TYPE "UDT012_Recirculation"
TITLE = State of recirculation mode
VERSION : 0.0
   STRUCT
      Intervall : Bool;   // Recirculation in interval mode (reduced or low pressure circulation)
      Parallel : Bool;   // Parallel circulation is activ (not used)
      Lowpressure : Bool;   // Low pressure circulation is active
      Reduced : Bool;   // Reduced circulation is active
      Highpressure : Bool;   // High pressure circulation over one mixing head is active
      Tolerance_OK : Bool;   // Request wether tolarances of the analog values at PUC are OK
      Weekendswitching : Bool;   // The pouring machine is in weekend mode
      Pausetime : Bool;   // The pouring machine is pausing time of the interval
      Break_KK : Bool;   // Stop flag of a active circulation mode to fill cylinder of a cylinder machine
      HP_is_active : Bool;   // High pressure circulation is active
      Is_selected : Bool;   // A circulation mode of the pouring machine is selected
      RequestPausePos : Bool;   // Request to the cylinder machine to bring the cylinder in break position
      cycle_runs : Bool;   // Save flag of the stop flag while starting a pouring cycle
      Is_active : Bool;   // A cycle mode of the pouring machine is active (no fault and oparition mode OK)
      Lowpressure_Exist : Bool;   // Low pressure circulation is existing
      Spare_1_7 : Bool;
      Switch_Intervall : Bool;   // Switch circulation in interval mode (reduced or low pressure circulation) selected
      Switch_Parallel : Bool;   // Switch Parallel circulation is selected (not used)
      Switch_Lowpressure : Bool;   // Switch Low pressure circulation is selected
      Switch_Reduced : Bool;   // Switch Reduced circulation is selected
      Intervall_Reduced : Bool;   // Reduced circulation in Intervall is active
      Intervall_Lowpressure : Bool;   // Low pressure circulation in Intervall is active
      Intervall_Reduced_Pause : Bool;   // Reduced circulation in Intervall pause is active
      Intervall_Lowpressure_Pause : Bool;   // Low pressure circulation in Intervall pause is active
      Spare_3_0 : Bool;
      Spare_3_1 : Bool;
      Spare_3_2 : Bool;
      Spare_3_3 : Bool;
      Spare_3_4 : Bool;
      Spare_3_5 : Bool;
      Spare_3_6 : Bool;
      Spare_3_7 : Bool;
      State_Intervall : Int;
      State_Lowpressure : Int;
      State_Reduced : Int;
      Indicator_HP : "UDT001_DWord_1_32";   // Indicates selected high pressure circulation
      Status_RC_HP : Int;   // Flag of the steps select and deselect high pressure circulation
      Button_HP : "UDT001_DWord_1_32";   // Button to select high pressure circulation
      Lamp_HP : "UDT001_DWord_1_32";   // Activation of lamps to indicat that high pressure recirculation runs
      SWU_RC_HP : DWord;   // Bitvalue of the SWU-Number where high pressure circulation runs
   END_STRUCT;
END_TYPE

TYPE "UDT013_Robot"
VERSION : 0.1
   STRUCT
      Switches : Struct
         SwitchHomePosON_OFF : Bool;   // Switch home position on/off
         SwitchMaintPosON_OFF : Bool;   // Switch maintenance position on/off
         SwitchTestShotON_OFF : Bool;   // Switch to make a couple shot with roboter
         SwitchCleaningON_OFF : Bool;   // Switch cleaning program on/off
         SwitchBrushON_OFF : Bool;   // Switch brush program on/off
         SwitchSyncON_OFF : Bool;   // Switch for checking EPS
         SwitchEnableRobotON_OFF : Bool;   // Switch no foaming in the conveyor (conveyor standalone)
         SwitchLearningON_OFF : Bool;   // Switch for learning the shot path (in conection with Shotware)
         SwitchTeachingON_OFF : Bool;   // Switch for Teaching the Robot
         Switch_10 : Bool;
         Switch_11 : Bool;
         Switch_12 : Bool;
         Switch_13 : Bool;
         Switch_14 : Bool;
         Switch_15 : Bool;
         Switch_16 : Bool;
         StateHomePos : Byte;   // 1->Drive ON; 2->Fault Drive; 3->Drive requested but not on
         StateMaintPos : Byte;   // 1->Drive ON; 2->Fault Drive; 3->Drive requested but not on
         StateTestShot : Byte;   // 1->Drive ON; 2->Fault Drive; 3->Drive requested but not on
         StateCleaning : Byte;   // 1->Drive ON; 2->Fault Drive; 3->Drive requested but not on
         StateBrush : Byte;   // 1->Drive ON; 2->Fault Drive; 3->Drive requested but not on
         StateSync : Byte;   // 1->Drive ON; 2->Fault Drive; 3->Drive requested but not on
         StateEnableRobot : Byte;   // 1->Drive ON; 2->Fault Drive; 3->Drive requested but not on
         StateLearning : Byte;   // 1->Drive ON; 2->Fault Drive; 3->Drive requested but not on
         StateTeaching : Byte;   // 1->Drive ON; 2->Fault Drive; 3->Drive requested but not on
         State_10 : Byte;
         State_11 : Byte;
         State_12 : Byte;
         State_13 : Byte;
         State_14 : Byte;
         State_15 : Byte;
         State_16 : Byte;
      END_STRUCT;
      State : Struct
         IRBInAuto : Bool;   // Robot in automatic
         IRBInManuel : Bool;   // Robot in manuel
         IRBtoHome : Bool;   // Robot to Homeposition
         IRBInHome : Bool;   // Robot in Homeposition
         IRBtoMaint : Bool;   // Robot to Maintenanceposition
         IRBInMaint : Bool;   // Robot in Maintenanceposition
         IRBtoClean : Bool;   // Robot to Cleaningposition
         IRBinClean : Bool;   // Robot in Cleaningposition
         IRBCleanEnd : Bool;   // Robot Cleaning finished
         IRBtoBrush : Bool;   // Robot to Brushposition
         IRBinBrush : Bool;   // Robot in Brushposition
         IRBCycleEnd : Bool;   // Robot Cycle end
         IRBOutRangeMC : Bool;   // Robot is out of the Mouldcarrier
         IRBError : Bool;   // Robot has an Error
         Reserve_12 : Bool;
         Reserve_13 : Bool;
         Reserve_14 : Bool;
         Reserve_15 : Bool;
         Reserve_16 : Bool;
         Reserve_17 : Bool;
         Reserve_18 : Bool;
         Reserve_19 : Bool;
         Reserve_20 : Bool;
         Reserve_21 : Bool;
         StepNumber : Byte;   // Stepnumber for stepchain of robot interface
      END_STRUCT;
   END_STRUCT;
END_TYPE

TYPE "UDT925_ShotResult"
VERSION : 0.1
   STRUCT
      PartNo : Int;   // Partnumber of shot at tool
      PartCounter : Int;
      FoamingTime : Real;   // Foaming Time
      PartWeight : Real;   // Part Weight
      Nitrogen : Real;   // Total value nitrogen from Inerting
      StationNo : Byte;
      Machine_No : Byte;
      MHNo : Byte := 0;   // Mixinghead number
      "Name" : Array[1..6] of String[20];
      Flow : Array[1..6] of Real;   // Flow for 8 components
      Pressure : Array[1..6] of Real;   // Pressure for 8 components
      Temperature : Array[1..6] of Real;   // Pressure for 8 components
      MaterialConsumption : Array[1..6] of Real;   // Flow for 8 components
      Mixingratio : Array[1..6] of Real;   // Flow for 8 components
      StausBitWarning : Array[1..6] of Struct
         StatusBitWarningMixingratio : Bool;
         StatusBitAlarmMixingratio : Bool;
         StatusBitWarningPressure : Bool;
         StatusBitAlarmPressure : Bool;
         StatusBitWarningPressureMH : Bool;
         StatusBitAlarmPressureMH : Bool;
         StatusBitWarningTemperature : Bool;
         StatusBitAlarmTemperature : Bool;
         StatusBitWarningTemperatureMH : Bool;
         StatusBitAlarmTemperatureMH : Bool;
         SpareBit11 : Bool;
         SpareBit12 : Bool;
         SpareBit13 : Bool;
         SpareBit14 : Bool;
         SpareBit15 : Bool;
         SpareBit16 : Bool;
      END_STRUCT;
      PartShotDisableService : Bool;
      StatusBitFaultGroup1 : Bool;
      StatusBitStopCycleDuringShot : Bool;
      ShotDisabledDuringShot : Bool;
      StatusBitManualShot : Bool;
      StatusBitAutomaticShot : Bool;   // Disable foaming
      SpareBit7 : Bool;   // Disable foaming
      SpareBit8 : Bool;   // Disable foaming
      StatusBitWarningFlow : Bool;
      StatusBitAlarmFlow : Bool;
      StatusBitWarningWeight : Bool;
      StatusBitAlarmWeight : Bool;
      StatusBitWarningFoamingTime : Bool;
      StatusBitAlarmFoamingTime : Bool;
      SpareBit15 : Bool;
      SpareBit16 : Bool;
   END_STRUCT;
END_TYPE

TYPE "UDT1810_Pentan"
VERSION : 0.1
   STRUCT
      FLT_PreAlarm_Pentan : Bool;
      FLT_PreAlam_NitrogenTank : Bool;
      FLT_NitrogenTank : Bool;
      FLT_Supply_Nitrogen : Bool;
      FLT_Exhausesystem : Bool;
      FLT_PentanpumpNotRunning : Bool;
      FLT_PentamixNotReady : Bool;
      MES_EStop_Pentamix : Bool;
      FLT_Valve1_Max : Bool;
      FLT_Valve2_Max : Bool;
      Spare_11 : Bool;
      Spare_12 : Bool;
      Spare_13 : Bool;
      Spare_14 : Bool;
      Spare_15 : Bool;
      Spare_16 : Bool;
   END_STRUCT;
END_TYPE

TYPE "UDT102_Pentan"
VERSION : 0.1
   STRUCT
      Fault_Exist : Bool;   // A fault inside this function exist
      FaultLevel_1 : Bool;   // A fault level 1 inside this function exist
      FaultLevel_2 : Bool;   // A fault level 2 inside this function exist
      FaultLevel_3 : Bool;   // A fault level 3 inside this function exist
      Message_Exist : Bool;   // A message inside this function exist
      EnableComponentPump : Bool;
      V_FillingValve1 : Bool;
      V_FillingValve2 : Bool;
      HM_Valve1_closed : Bool;
      HM_Valve2_closed : Bool;
      HM_FillingValve1 : Bool;
      HM_FillingValve2 : Bool;
      HM_FillingValve1_Opened : Bool;
      HM_FillingValve2_Opened : Bool;
      HMFillingValves_Open : Bool;
      HM_FillingValve : Bool;
   END_STRUCT;
END_TYPE

TYPE "UDT780_ParaPW_Controller"
VERSION : 0.1
   STRUCT
      Max_Temp_Diff_Cooling : Real;   // Maximum difference of Temperature cooling
      Max_Temp_Diff_Heating : Real;   // Maximum difference of Temperature heating
      PLC_Control_Area : Real;   // time
      Weighting_Temp : Real;   // Weighting of two temperatures
      Offset_Cooling : Real;
      Offset_Heating : Real;
   END_STRUCT;
END_TYPE

TYPE "UDT106_ControllerHeatExchanger"
TITLE = State of 2-point controller tempering
VERSION : 0.1
   STRUCT
      CoolingActive : Bool;
      HeatingActive : Bool;
      CoolingRequest : Bool;
      HeatingRequest : Bool;
      FLT_Fuse_Heating : Bool;
      HF_Set_Cooling : Bool;
      HF_Set_Heating : Bool;
      Spare_13 : Bool;
      Trigger : Bool;   // Trigger to start calculation pulstime
      Start_delay_puls : Bool;
      Fault_Exist : Bool;
      Spare_1_3 : Bool;
      Spare_1_4 : Bool;
      Spare_1_5 : Bool;
      Spare_1_6 : Bool;
      Switch_Temp_ON_OFF : Bool;
      PulsTime : Real;   // Time to switch on valve heatexchanger
      State_Temp : Int;
   END_STRUCT;
END_TYPE

TYPE "UDT124_Inerting"
VERSION : 0.1
   STRUCT
      FaultLevel_1 : Bool;   // A fault group 1 exist
      FaultLevel_2 : Bool;   // A fault group 2 exist
      FaultLevel_3 : Bool;   // A fault group 3 exist
      Message_activ : Bool;   // A message is active
      Reserve14 : Bool;
      Reserve15 : Bool;
      Reserve16 : Bool;
      Reserve17 : Bool;
      OK : Bool;   // Inerting finished
      Inert_canceled : Bool;   // Inerting canceled
      Start_PressurizeTimeRuns : Bool;   // Start pressureize time
      Inert_runs : Bool;   // Inerting runs
      Inert_started : Bool;   // Waiting for shottime
      Purge_runs : Bool;   // Purge mixhead is activ
      Inert_ON_OFF : Bool;   // Inerting on/off over refernce value
      Inert_Off_Dry_Shot : Bool;   // Inerting off for dry shot
      FH_Start : Bool;
      FP_Start : Bool;
      FH_ST_received : Bool;
      FP_ST_received : Bool;   // Shottime received
      FH_Stop : Bool;
      FP_Stop : Bool;   // Stop cycle if fault
      Set_LoadValue : Bool;
      Reserve27 : Bool;
      FH_Start_Time : Bool;
      FP_Start_Time : Bool;
      FP_Start_Inert : Bool;
      FH_Start_Inert : Bool;
      FP_Start_Leakage_Control : Bool;
      FH_Start_Leakage_Control : Bool;
      Reserve26 : Bool;
      Reserve28 : Bool;
      FN_CP_after_Shot : Bool;
      FN_Prepare_Purge_after_Shot : Bool;
      Start_Prepare_Purge_after_Shot : Bool;
      Start_Purge_after_Shot : Bool;
      Start_Purge_Manual : Bool;
      HF_Start_Purge_Manual : Bool;
      Enable_Purge : Bool;
      FN_Purge_after_shot_finished : Bool;
      Reserve40 : Bool;
      Reserve41 : Bool;
      Reserve42 : Bool;
      Reserve43 : Bool;
      Reserve44 : Bool;
      Reserve45 : Bool;
      Reserve46 : Bool;
      Reserve47 : Bool;
      Purge_after_Shot : S5Time := S5T#400MS;
      Computed_Value : Real;
      Actual_Flow_N2 : Real;
      Actual_Flow_N2_measured_Total : Real;
      Actual_Flow_N2_Visu : Real;
      Total_Flow_N2_Visu : Real;
      Leakage_Actual_Flow_N2_measured_Total : Real;
      Leakage_Actual_Flow_N2_Visu : Real;
      Leakage_Total_Flow_N2_Visu : Real;
   END_STRUCT;
END_TYPE

TYPE "UDT125_Inerting_SetValues"
VERSION : 0.1
   STRUCT
      with_Purge : Bool;
      with_purge_after_Shot : Bool;
      with_Interval_Purge : Bool;
      with_Cycle_before_Inert_finished : Bool;
      with_inert_over_MH : Bool;
      with_inert_over_Lance : Bool;
      with_output_without_N2 : Bool;
      Inert_Switch_ON_OFF : Bool;
      Reservebyte : Byte;
      Reference_Value_Inert : Real := 0.0;
      Max_Reference_Value_Inert : Real;
      Foam_density : DInt := 350;
      Inerting_factor : Real := 10.0;
      Start_Offset : Real;
      Leakage_Value : Real;
      Reserve1 : Real;
      Inerting_time : S5Time;
      Max_Inerting_Time : S5Time := S5T#30S;
      Ready_Time_after_Inert : S5Time := S5T#10S;   // Reserve 245
      Delay_Plunger : S5Time := S5T#2S;   // Reserve 189
      Delay_Purge : S5Time := S5T#2S;
      Purge_time : S5Time := S5T#1S;
      Purge_after_Shot : S5Time := S5T#400MS;
      Delay_Purge_Interval : S5Time;
      Purge_Time_interval : S5Time;
      Pause_Time_interval : S5Time;
      Duration_Time_Interval : S5Time;
      Reserve2 : S5Time;
      Reserve3 : S5Time;
      Reserve4 : S5Time;
   END_STRUCT;
END_TYPE

TYPE "UDT021_Hydr_State"
TITLE = State of hydraulic
VERSION : 0.0
   STRUCT
      Switch_on_Motor : Bool;   // Release switch hydraulic motor on (feedback)
      MH_Hyd_OK : Bool;   // Hydraulic runs and operation pressure is reached
      Startup_Motor_finished : Bool;   // Start up hydraulic motors finished
      Switch_Hydraulic_ON_OFF : Bool;   // Switch ON/OFF hydraulic motor (external signal)
      FaultLevel_1 : Bool;   // A fault group 1 exist
      FaultLevel_2 : Bool;   // A fault group 2 exist
      FaultLevel_3 : Bool;   // A fault group 3 exist
      Fault_Exist : Bool;   // An actual fault exist
      Spare_09 : Bool;   // There is a mainfault -> hydraulic motor stopped
      Request_from_CP : Bool;   // Request from cleaning piston to build up hydraulic pressure
      Act_PressureBuildUp : Bool;   // Activation of the pressure build up valve
      Act_Main : Bool;   // Activation of mains contacor hydraulik- motor
      Act_Star : Bool;   // Activation of star contacor hydraulik- motor
      Act_Delta : Bool;   // Activation of delta contacor hydraulik- motor
      Act_Oilcooling : Bool;   // Activation of the oil cooling valve
      Spare_16 : Bool;
      State_Hydraulic : Int;   // 1->Drive ON; 2->Fault Drive; 3->Drive requested but not on
      HourCounter : DInt := 0;   // Hour counter of mixinghead hydraulic
   END_STRUCT;
END_TYPE

TYPE "UDT022_Zyl_Hyd_State"
TITLE = State of piston hydraulic
VERSION : 0.0
   STRUCT
      Request_Motor : Bool;   // Switch ON Hydraulic motor
      Hyd_ok : Bool;   // Hadraulic start up finished
      Fault_Min_Level : Bool;   // Fault: min level hydraulic oil
      WRN_C_Max : Bool;   // Warning: max temperature hydraulic oil
      Fault_C_Max : Bool;   // Fault: Maximum temperature of hydraulic oil was exceeded more than 5 minutes
      Fault_Motorprotection : Bool;   // Fault: Motorprotection hydraulic drive motor
      Fault_Filter : Bool;   // Fault: filter hydraulic is polluted
      Fault_Moog_Filter : Bool;   // Fault: Pre run high pressure filter is polluted
      mains_contactor : Bool;   // Activation of mains contacor hydraulik- motor
      Star_contactor : Bool;   // Activation of star contacor hydraulik- motor
      Delta_contactor : Bool;   // Activation of delta contacor hydraulik- motor
      FaultLevel_1 : Bool;   // A fault group 1 exist
      FaultLevel_2 : Bool;   // A fault group 2 exist
      FaultLevel_3 : Bool;   // A fault group 3 exist
      Reserve_1_6 : Bool;
      Programblock_is_active : Bool;   // Function block is active // Info at least 1 piston is active
   END_STRUCT;
END_TYPE

TYPE "UDT1825_FLT_Inerting"
VERSION : 0.1
   STRUCT
      Sensor_FLT_broken_wire : Bool;   // There is no connection to the sensor (3)
      Warning_limit_plus : Bool;   // The lower warning limit of the processvalue under run (3)
      Warning_limit_minus : Bool;   // The upper warning limit of the processvalue is exceeded (3)
      Alarm_limit_plus : Bool;   // The lower alarm limit of the processvalue under run(1)
      Alarm_limit_minus : Bool;   // The upper alarm limit of the processvalue is exceeded (1)
      Controller_at_limit : Bool;   // Controller at limit (3)
      Reserve1 : Bool;
      Fuse_TemperingOverLoad : Bool;   // Circuit breaker fault
      Fault_P_N2 : Bool;   // Fault Nitrogen Pressure
      Fault_flow_N2 : Bool;   // Fault Nitrogen Flowrate
      Fault_P_Flushing_Agent : Bool;   // Fault Flushing Agent
      Fault_Leakage_N2 : Bool;   // Fault Leakage Nitrogen
      Fault_MaxInertingTime : Bool;   // Maximum time for inerting
      Fault_NoShotwight : Bool;   // No shotwight or program number 0 or over 99
      Reserve16 : Bool;
      Reserve17 : Bool;
   END_STRUCT;
END_TYPE

TYPE "UDT126_Inerting_ActValues_Ma"
VERSION : 0.1
   STRUCT
      Actual_Flow_N2 : Real;
      Actual_Flow_N2_measured_Total : Real;
      Actual_Flow_N2_Visu : Real;
      Total_Flow_N2_Visu : Real;
      Leakage_Actual_Flow_N2_measured_Total : Real;
      Leakage_Actual_Flow_N2_Visu : Real;
      Leakage_Total_Flow_N2_Visu : Real;
   END_STRUCT;
END_TYPE

TYPE "Kuka_KRC4_Input"
VERSION : 0.1
   STRUCT
      E_KRC_STOPMES : Bool;   // Störmeldung aufgetreten
      E_KRC_PGNO_REQ : Bool;   // Programmnummer übermitteln
      E_KRC_APPL_RUN : Bool;   // Ein Programm wird abgearbeitet
      E_KRC_PERI_RDY : Bool;   // Antriebe sind eingeschaltet
      E_KRC_ALARM_STOP : Bool;   // Not-Halt aufgetreten
      E_KRC_USER_SAF : Bool;   // Schutzgitter / Zustimmschalter offen
      E_KRC_T1 : Bool;   // Betriebsart T1 am Schäumroboter angewählt
      E_KRC_T2 : Bool;   // Betriebsart T2 am Schäumroboter angewählt
      E_KRC_AUT : Bool;   // Betriebsart Automatik am Schäumroboter angewählt
      E_KRC_AUT_EXTERN : Bool;   // Betriebsart Automatik extern am Schäumroboter angewählt
      E_KRC_ON_PATH : Bool;   // Schäumroboter befindet sich auf der programmierten Bahn
      E_KRC_PRO_ACT : Bool;   // Roboter Prozess aktiv
      E_KRC_IN_HOME : Bool;   // Schäumroboter in Homeposition
      E_KRC_RC_READY : Bool;   // Fehler in der Robotersteuerung
      E_KRC_MH_in_FoamPos : Bool;   // MK ist in Schäumposition
      E_KRC_Blowair : Bool;   // Signal zum Ausblasen des MK
      E_KRC_FLT_WaitTime : Bool;
      E_KRC_IN_MAINPOS : Bool;   // Roboter ist in Wartungsposition
      E_KRC_OUT_19 : Bool;
      E_KRC_OUT_20 : Bool;
      E_KRC_OUT_21 : Bool;
      E_KRC_OUT_22 : Bool;
      E_KRC_IN_CLEANPOS : Bool;   // Roboter ist in Reinigungsposition
      E_KRC_MH_OPEN : Bool;   // Roboter ist in Schäumposition (PU kann Mischkopf öffnen)
      E_KRC_FOAMPROG_FINISHED : Bool;   // Roboter meldet alle Schüsse Schäumprogramm beendet
      E_KRC_OUT_26 : Bool;
      E_KRC_OUT_27 : Bool;
      E_KRC_OUT_28 : Bool;
      E_KRC_OUT_29 : Bool;
      E_KRC_OUT_30 : Bool;
      E_KRC_OUT_31 : Bool;
      E_KRC_OUT_32 : Bool;
      E_KRC_OUT_33 : Bool;
      E_KRC_OUT_34 : Bool;
      E_KRC_OUT_35 : Bool;
      E_KRC_OUT_36 : Bool;
      E_KRC_OUT_37 : Bool;
      E_KRC_OUT_38 : Bool;
      E_KRC_OUT_39 : Bool;
      E_KRC_OUT_40 : Bool;
      E_KRC_OUT_41 : Bool;
      E_KRC_OUT_42 : Bool;
      E_KRC_OUT_43 : Bool;
      E_KRC_OUT_44 : Bool;
      E_KRC_OUT_45 : Bool;
      E_KRC_OUT_46 : Bool;
      E_KRC_OUT_47 : Bool;
      E_KRC_OUT_48 : Bool;
   END_STRUCT;
END_TYPE

TYPE "Fanuc_Input"
VERSION : 0.1
   STRUCT
      Robi_stop_extern : Bool;   // 1:UI1 (0) - immediate stop (sofortiger Halt) -> Not Aus
      HOLD_to_Robot : Bool;   // 2:UI2 (0) - Roboter bremst bis zum stillstand ab, Programm wird angehalten
      Robot_safety_speed : Bool;   // 3:UI3 (0) - Sicherheitsgeschwindigkeit -> Anhalten des Robo bei Sicherhei niO
      CSTOPI_to_Robot : Bool;   // 4:UI4 (0) - Cycle stop -> Beendung des Programm nach der Ausführung
      Robot_Fault_reset : Bool;   // 5:UI5 (1) - Einschalten der Servospannung -> Alarm quittieren
      START_Robot : Bool;   // 6:UI6 (1) - Zum Starten der bereits abgebrochemem Ablaufprogramme
      Move_to_home_to_Robot : Bool;   // 7:UI7 (1) -
      Enable_Robi_SPS_RN : Bool;   // 8:UI8 (1) - Aktivierungssignal -> Freigabe zur Bewegung
      PNS01 : Bool;   // 9:UI9 (1) - Aufruf des Ablaufprogrammes
      PNS02 : Bool;   // 10:UI10 (1) - Aufruf des Ablaufprogrammes
      PNS03 : Bool;   // 11:UI11 (1) - Aufruf des Ablaufprogrammes
      PNS04 : Bool;   // 12:UI12 (1) - Aufruf des Ablaufprogrammes
      PNS05 : Bool;   // 13:UI13 (1) - Aufruf des Ablaufprogrammes
      PNS06 : Bool;   // 14:UI14 (1) - Aufruf des Ablaufprogrammes
      PNS07 : Bool;   // 15:UI15 (1) - Aufruf des Ablaufprogrammes
      PNS08 : Bool;   // 16:UI16 (1) - Aufruf des Ablaufprogrammes
      PNS_STROBE_to_Robot : Bool;   // 17:UI17 (1) - Zum Starten der Auswahl der ainzelnen Ablaufprogramme
      PROD_START_to_Robot : Bool;   // 18:UI18 (1) - Zum Starten der einzelnen Ablaufprogramme
      di01_1 : Bool;   // 19/1:
      di01_2 : Bool;   // 20/2:
      di01_3 : Bool;   // 21/3:
      di01_4 : Bool;   // 22/4:
      di01_5 : Bool;   // 23/5:
      di01_6 : Bool;   // 24/6:
      di01_7 : Bool;   // 25/7:
      di01_8 : Bool;   // 26/8:
      di01_9 : Bool;   // 27/9:
      di01_10 : Bool;   // 28/10:
      di01_11 : Bool;   // 29/11:
      diSync : Bool;   // 30/12:
      diBreak : Bool;   // 31/13:Signal zum auslösen des Interrupt 1 // Programm stoppen
      diInterrupt : Bool;   // 32/14:Signal zum auslösen des Interrupt 2
      diStartCycle : Bool;   // 33/15:Signal to start the robotcycle
      diReadProgNo : Bool;   // 34/16:A programnumber can read from PLC
      diRelMoveMC : Bool;   // 35/17:The robot can start with it´s movements
      diShotDigIn : Bool;   // 36/18:Spare
      diStartCleanMH : Bool;   // 37/19:The robot can move to MH-Cleaningstation
      diCleanMHEnd : Bool;   // 38/20:The MH-Cleaning is finished
      diStartBrushMH : Bool;   // 39/21:The robot can move to the brush station
      diHomeToPreP : Bool;   // 40/22:Spare
      diHomeToMaintP : Bool;   // 41/23:Signal to move the robot from homeposition to maintenanceposition
      diMaintToHomeP : Bool;   // 42/24:Signal to move the robot from maintenanceposition to homeposition
      diRobinSafepos : Bool;   // 43/25:Signal that the other robot is in a safe position
      diProgBreak : Bool;   // 44/26:Signal to break the program
      diJumpConveyor : Bool;   // 45/27:Spare
      diBackToRest : Bool;   // 46/28:Signal to move the robot back to homeposition after foaming
      diEnblNextMould : Bool;   // 47/29:Freigabe zum Fahren in die nächste Form
      diEnableHome : Bool;   // 48/30: Enable signal for movement to home position (other robot is in home)
      diPLCWaitWobj : Bool;   // 49/31:Signal to activate the waitwobj instruction
      diPLCDropWobj : Bool;   // 50/32:Signal to drop the activ wobj
      diSingleOP : Bool;   // 51/33:Signal for emergency production with this robot only
      diMC_is_open : Bool;   // 52/34:
      diLoad_MC : Bool;   // 53/35:
      diMove_out_MC : Bool;   // 54/36:
      diQuickStop : Bool;   // 55/37:
      diRel2ndMould : Bool;   // 56/38: Conv. Position ok to shift in 2n mould
      diBolt1 : Bool;   // 57/39:
      diBolt2 : Bool;   // 58/40:
      diGripper_stretched : Bool;   // 59/41:
      diGripper_unstretched : Bool;   // 60/42:
      diGripper_open : Bool;   // 61/43:
      diGripper_closed : Bool;   // 62/44:
      diEnblClosingArea : Bool;   // 63/45:
      diSyncConveyor : Bool;   // 64/46:
      diBlockInitOrgtrigger : Bool;   // 65/47: Block the ORGTRIGGER init because of teaching Robot 2
      diHomeToTestP : Bool;   // 66/48: Signal to move the robot from homeposition to test shot position
      diTestToHomeP : Bool;   // 67/49: Signal to move the robot from test shot position to home position
      diAction_04 : Bool;   // 68/50:Action 4 activ
      diAction_05 : Bool;   // 69/51:Action 5 activ
      diAction_06 : Bool;   // 70/52:Action 6 activ
      diAction_07 : Bool;   // 71/53:Action 7 activ
      diAction_08 : Bool;   // 72/54:Action 8 activ
      diAction_09 : Bool;   // 73/55:Action 9 activ
      diAction_10 : Bool;   // 74/56:Action 10 activ
      di10_57 : Bool;   // 75/57:Spare
      di10_58 : Bool;   // 76/58:Spare
      di10_59 : Bool;   // 77/59:Spare
      di10_60 : Bool;   // 78/60:Spare
      di10_61 : Bool;   // 79/61:Spare
      di10_62 : Bool;   // 80/62:Spare
      giMouldCodeBit0 : Bool;   // 81/63:Anzahl der Formen im Formträger (Gruppeingang Bit 0)
      giMouldCodeBit1 : Bool;   // 82/64:Anzahl der Formen im Formträger (Gruppeingang Bit 1)
      di01_065 : Bool;   // 83/65:
      di01_066 : Bool;   // 84/66:
      di01_067 : Bool;   // 85/67:
      di01_068 : Bool;   // 86/68:
      di01_069 : Bool;   // 87/69:
      di01_070_SyncTest : Bool;   // 88/70:
      GIMCNo : Byte;   // 89/71:Nummer des Formträgers der Form// Abhängig vom MouldCode
      GIProgNo1 : Int;   // 97/79:Verfahrprogramm für die erste Form // Eingetragen in PUC
      GIProgNo2 : Int;   // 113/95:Verfahrprogramm für die zweite Form // Eingetragen in PUC
      giTeachProgNo1 : Int;   // 129/111: Verfahrprogramm für die erste Form zum Teachen
      giTeachProgNo2 : Int;   // 145/127: Verfahrprogramm für die zweite Form zum Teachen
   END_STRUCT;
END_TYPE

TYPE "Kuka_KRC4_Status"
VERSION : 0.1
   STRUCT
      STG_System : Bool;
      STG_Schnittstelle : Bool;
      STG_Roboter_stoppt : Bool;
      STG_Motoschutz : Bool;
      STG_0_4 : Bool;
      STG_0_5 : Bool;
      STG_0_6 : Bool;
      STG_0_7 : Bool;
      STG_0_8 : Bool;
      STG_0_9 : Bool;
      STG_0_10 : Bool;
      STG_0_11 : Bool;
      STG_0_12 : Bool;
      STG_0_13 : Bool;
      STG_0_14 : Bool;
      STG_0_15 : Bool;
      Anforderung_MP : Bool;
      Anforderung_Reinigen : Bool;
      PrgNr_ok : Bool;
      HM_Ext_Start : Bool;
      FHM_PrgNr_gueltig : Bool;
      FHM_PRG_laeuft : Bool;
      FHM_FRG_schaeumen : Bool;
      FRG_schaeumen : Bool;
      FHM_PRO_ACT : Bool;
      Anforderung_Automatik : Bool;
      Warten_auf_MK_Reinigung : Bool;
      FHM_Teischuss_Null : Bool;
      FHM_MainPosToHomePos : Bool;
      FHM_HomePosToMainPos : Bool;
      FHM_Cleaning_MH : Bool;
      Spare_4 : Bool;
      Spare_5 : Bool;
      Spare_6 : Bool;
      Spare_7 : Bool;
      Spare_8 : Bool;
      Spare_9 : Bool;
      Spare_10 : Bool;
      Spare_11 : Bool;
      Spare_12 : Bool;
      Spare_13 : Bool;
      Spare_14 : Bool;
      Spare_15 : Bool;
      Spare_16 : Bool;
      Spare_17 : Bool;
      A_SPS_PGNO : Byte;
      SpareDint_1 : DInt;
      SpareDint_2 : DInt;
      SpareDint_3 : DInt;
      SpareDint_4 : DInt;
      Input_From_Robot : "Kuka_KRC4_Input";
      Output_To_Robot : "Kuka_KRC4_Output";
   END_STRUCT;
END_TYPE

TYPE "Fanuc_Output"
VERSION : 0.1
   STRUCT
      CMDENBL_Robot_ready : Bool;   // 1:UO1 - Die Remote Bedingungen sind erfüllt (Roboter bereit)
      SYSRDY_Robot_sys_ready : Bool;   // 2:UO2 - Die Servospannung ist eingeschaltet -> Rooboter bereit
      Robot_Prgrun : Bool;   // 3:UO3 - Programm läuft, wird ausgeführt
      Robot_Prg_paused : Bool;   // 4:UO4 - Programm wurde unterbrochen -> wartet auf Neustart
      Robot_motion_held : Bool;   // 5:UO5 - HOLD- Taste ist betätigt
      Fault_Robot : Bool;   // 6:UO6 - Alarm steht an
      Robot_at_home_Pos : Bool;   // 7:UO7 - Roboter in Refernezposition -> Hier Homeposition
      Robot_TP_enabled : Bool;   // 8:UO8 - Der Aktivierungsschalter am Teachpanel wird betätigt
      Robot_Batt_alarm : Bool;   // 9:UO9 - Die Spannung an der Backup- Battery ist zu niedrig
      Robot_busy : Bool;   // 10:UO10 - Ein Programm/ Prozedure läuft, wird ausgeführt
      SNO01 : Bool;   // 11:UO11 - Ausgabe des aktuellen Programms
      SNO02 : Bool;   // 12:UO12 - Ausgabe des aktuellen Programms
      SNO03 : Bool;   // 13:UO13 - Ausgabe des aktuellen Programms
      SNO04 : Bool;   // 14:UO14 - Ausgabe des aktuellen Programms
      SNO05 : Bool;   // 15:UO15 - Ausgabe des aktuellen Programms
      SNO06 : Bool;   // 16:UO16 - Ausgabe des aktuellen Programms
      SNO07 : Bool;   // 17:UO17 - Ausgabe des aktuellen Programms
      SNO08 : Bool;   // 18:UO18 - Ausgabe des aktuellen Programms
      ROB_SNACK_Prg_valid : Bool;   // 19:UO19 - Programm wurde angenommen
      UO020 : Bool;   // 20:UO20 - Reserve
      do_IRB_Auto : Bool;   // 21/1:Schlüsselschalter am Roboter auf Automatik- Betrieb
      do_IRB_Manual_20 : Bool;   // 22/2:Schlüsselschalter am Roboter auf Hand 20%- Betrieb
      do_IRB_Manual_100 : Bool;   // 23/3:3chlüsselschalter am Roboter auf Hand 100%- Betrieb
      doEmStop_Akt : Bool;   // 24/4:Robot is in Status Emergency Stop
      doIRBInHome : Bool;   // 25/5:Der Roboter befindet sich in seiner Grundposition
      doIRBInMaintP : Bool;   // 26/6:Der Roboter befindet sich in seiner Wartungsposition
      doIRBOutRange : Bool;   // 27/7:Der Roboter befindet sich in der Nähe seines Arbeitsbereiches
      doIRBOutRangemc : Bool;   // 28/8:Der Roboter befindet sich außerhalb des Störbereiches des Formträgers
      do01_9 : Bool;   // 29/9:
      do01_10 : Bool;   // 30/10:
      do01_11 : Bool;   // 31/11:
      do01_12 : Bool;   // 32/12:
      doCycleStarted : Bool;   // 33/13:The programcycle is startet
      doCycleEnd : Bool;   // 34/14:The programcycle is finished
      doProgNoRead : Bool;   // 35/15The programnumber is readed
      doShotDigOut : Bool;   // 36/16:1'ter digitaler Ausgang der Shotware // Mischkopf öffnen
      doStopFoamPLC : Bool;   // 37/17:Signal to stop the foaming because the robotprogram has stoped
      doCloseMouldF : Bool;   // 38/18:Signal that the robot is out of the mould
      doCleaningPLC : Bool;   // 39/19:Ansteuererung eines Mischkopfreinigers oder des Reinigungskolben
      doIRBSyncWobj : Bool;   // 40/20:Der Roboter wurde aufsyncronisiert (Tracking)
      doRobWaitWobj : Bool;   // 41/21:Der Roboter wartet auf das aufsyncronisieren (Tracking)
      doCleanOsziJet : Bool;   // 42/22:Ansteuerung der Luft zum Freibl. von Oszillierdüsen bei Faseransteuerung
      doBlowAir : Bool;   // 43/23:Ansteuerung der Blasluft im Mischkopf bei einer Faseransteuerung
      doCleanBrushOn : Bool;   // 44/24:Ansteuerung einer Einrichtung zum reinigen des Mischkopfes
      doShotDigOut2 : Bool;   // 45/25:2'ter digitaler Ausgang der Shotware // Längenverstellung
      doInPosTeach : Bool;   // 46/26:Der Roboter befindet sich in der Position zum Teachen
      doConveyorStoped : Bool;   // 47/27:Der Conveyor steht// Impulseingänge werden nicht erkannt
      doReadyToStart : Bool;   // 48/28:Der Roboter ist fertig für den gemeinsamen Start mehrerer Roboter
      doBackToRest : Bool;   // 49/29:Roboter ist fertig für die gemeinsame Bewegung zur Homeposition
      doRPELoading : Bool;   // 50/30:SONDER für Johnson Controlls: RPE Module werden geladen
      doErrLoadMoRPE : Bool;   // 51/31:SONDER für Johnson Controlls: RPE Fehler beim Module laden
      doFlushing : Bool;   // 52/32:
      doHornLuft : Bool;   // 53/33:
      doZerstaeuberLuft : Bool;   // 54/34:
      doSpuelen_1 : Bool;   // 55/35:
      doSpuelen_2 : Bool;   // 56/36:
      doBolt1 : Bool;   // 57/37:
      doBolt2 : Bool;   // 58/38:
      doIRBInTestP : Bool;   // 59/39: Der Roboter befindet sich in der Testschussposition
      doNoValidPrg : Bool;   // 60/40: No valid program number found
      do01_041 : Bool;   // 61/41:
      do01_042 : Bool;   // 62/42:
      do01_043 : Bool;   // 63/43:
      do01_044 : Bool;   // 64/44:
      doAction_01 : Bool;   // 65/45:Action 01 activ
      doAction_02 : Bool;   // 66/46:Action 02 activ
      doAction_03 : Bool;   // 67/47:Action 03 activ
      doAction_04 : Bool;   // 68/48:Action 04 activ
      doAction_05 : Bool;   // 69/49:Action 05 activ
      doAction_06 : Bool;   // 70/50:Action 06 activ
      doAction_07 : Bool;   // 71/51:Action 07 activ
      doAction_08 : Bool;   // 72/52:Action 08 activ
      doAction_09 : Bool;   // 73/53:Action 09 activ
      doAction_10 : Bool;   // 74/54:Action 10 activ
      do10_55 : Bool;   // 75/55:Reserve
      do10_56 : Bool;   // 76/56:Reserve
      do10_57 : Bool;   // 77/57:Reserve
      do10_58 : Bool;   // 78/58:Reserve
      do10_59 : Bool;   // 79/59:Reserve
      do10_60 : Bool;   // 80/60:Reserve
      do01_61_77 : Word;   // 81/61:
      GO_Reserve : Byte;   // 97/77:
      goFormAktBit0 : Bool;   // 105/85:Nummer der Form (1.3) welche zur Zeit bearbeitet wird (Gruppenausgang 0)
      goFormAktBit1 : Bool;   // 106/86:Nummer der Form (1.3) welche zur Zeit bearbeitet wird (Gruppenausgang 1)
      go01_087 : Bool;   // 107/87:
      go01_088 : Bool;   // 108/88:
      go01_089 : Bool;   // 109/89:
      go01_090 : Bool;   // 110/90:
      go01_091 : Bool;   // 111/91:
      go01_092 : Bool;   // 112/92:
      GOError : Byte;   // 113/93:Fehlernummer bei der Bearbeitung des Programms (Gruppenausgang)
      go01_101_109 : Byte;   // 121/101:
      goxFIProgBit0 : Bool;   // 129/109:Nummer des Faserprogrammes an PUC (Gruppenausgang der Shotware, Bit 0)
      goxFIProgBit1 : Bool;   // 130/110:Nummer des Faserprogrammes an PUC (Gruppenausgang der Shotware, Bit 1)
      goxFIProgBit2 : Bool;   // 131/111:Nummer des Faserprogrammes an PUC (Gruppenausgang der Shotware, Bit 2)
      goxFIProgBit3 : Bool;   // 132/112:Nummer des Faserprogrammes an PUC (Gruppenausgang der Shotware, Bit 3)
      go01_113 : Bool;   // 133/113:
      go01_114 : Bool;   // 134/114:
      go01_115 : Bool;   // 135/115:
      go01_116 : Bool;   // 136/116:
      goOscixFIBit0 : Bool;   // 137/117:Bit des Oszillierprogrammes // X1 (2'ter GroupOut der Shotware, Bit 0)
      goOscixFIBit1 : Bool;   // 138/118:Bit des Oszillierprogrammes // X2 (2'ter GroupOutder Shotware, Bit 1)
      goOscixFIBit2 : Bool;   // 139/119:Bit des Oszillierprogrammes // Y1 (2'ter GroupOut der Shotware, Bit 2)
      goOscixFIBit3 : Bool;   // 140/120:Bit des Oszillierprogrammes // Y2 (2'ter GroupOut der Shotware, Bit 3)
      go01_121 : Bool;   // 141/121:
      go01_122 : Bool;   // 142/122:
      go01_123 : Bool;   // 143/123:
      go01_124 : Bool;   // 144/124:
      goReserveXX : Word;   // 145/125:
   END_STRUCT;
END_TYPE

TYPE "Kuka_KRC4_Output"
VERSION : 0.1
   STRUCT
      A_SPS_PGNO : Byte;   // Programmnummer an den Schäumroboter
      A_SPS_PARITY : Bool;   // Paritäts-Bit der Programmnummer
      A_SPS_PGNO_VALID : Bool;   // Programmnummer einlesen
      A_SPS_EXT_START : Bool;   // Programm Start
      A_SPS_MOVE_ENABLE : Bool;   // Antriebsfreigabe Roboter
      A_SPS_CONF_MESS : Bool;   // Fehlermeldung extern quitt.
      A_SPS_DRIVES_ON : Bool;   // Antriebe einschalten
      A_SPS_DRIVES_OFF : Bool;   // Antriebe auschalten
      A_KRC_MOVE_TO_HOMEPOS : Bool;   // Roboter soll in die Homeposition fahren
      A_KRC_MOVE_TO_CLEANPOS : Bool;   // Roboter soll in die Reinigungsposition fahren
      A_KRC_MOVE_TO_MAINPOS : Bool;   // Roboter soll in die Wartungsposition fahren
      A_SPS_DIRELMOVEMC : Bool;   // Freigabe für Bewegung in die Form
      A_KRC_IN_20 : Bool;
      A_KRC_IN_21 : Bool;
      A_KRC_IN_22 : Bool;
      A_SPS_PU_OK : Bool;   // PU in Automatikbetrieb und OK
      A_SPS_CYCLE_RUN : Bool;   // Zyklus läuft (Maschine baut Druck auf)
      A_SPS_READY_FOR_SHOT : Bool;   // Schussbereit (Maschine ist bereit zum Schuss)
      A_SPS_SHOT_RUNS : Bool;   // Schuss läuft
      A_SPS_SHOTEND : Bool;   // Schussende
      A_SPS_SERVICE : Bool;   // Service (Simulationsbetrieb/Trockenschuss)
      A_SPS_INTERRUPT : Bool;   // Abbruch
      A_KRC_IN_30 : Bool;
      A_KRC_IN_31 : Bool;
      A_KRC_IN_32 : Bool;
      A_KRC_IN_33 : Bool;
      A_KRC_IN_34 : Bool;
      A_KRC_IN_35 : Bool;
      A_KRC_IN_36 : Bool;
      A_KRC_IN_37 : Bool;
      A_KRC_IN_38 : Bool;
      A_KRC_IN_39 : Bool;
      A_KRC_IN_40 : Bool;
      A_KRC_IN_41 : Bool;
      A_KRC_IN_42 : Bool;
      A_KRC_IN_43 : Bool;
      A_KRC_IN_44 : Bool;
      A_KRC_IN_45 : Bool;
      A_KRC_IN_46 : Bool;
      A_KRC_IN_47 : Bool;
      A_KRC_IN_48 : Bool;
   END_STRUCT;
END_TYPE

TYPE "UDT_TT_SafetyDevice"
VERSION : 0.1
   STRUCT
      OpeningSelected : Bool;   // Opening of the safety device is selected
      OpeningEnabled : Bool;   // Opening of the safety device is possible
      EdgeButton : Bool;   // Edge of the button to select opening of the safety device
      HFEdgeButton : Bool;   // Help flag for the edge
      EdgeASReset : Bool;   // Edgo of the reset of Auto Stop from this safety device
      HFEdgeASReset : Bool;   // Help flag for the edge
      HFforMESSelected : Bool;   // Help flag for the message opening is selected
      HFforMESAutomaticStop : Bool;   // Help flag for message automatic stop is activ
      Spare1 : Byte;
   END_STRUCT;
END_TYPE

TYPE "General_Faults"
VERSION : 0.1
   STRUCT
      FLT_System : Bool;   // System fault from robot
      FLT_Interface : Bool;   // Interface faulty
      FLT_Prog_stopped : Bool;   // Rob prog stopped
      FLT_Fuse : Bool;   // Fault fuse
      FLT_Wrong_Prog_No : Bool;   // Prog no. not existing
      FLT_Wrong_MC_No : Bool;   // Workobject not existing
      FLT_Wrong_Shot_time : Bool;   // Shot time too short (Shotware)
      FLT_TP_On_in_automatic : Bool;   // TP is ON in automatic mode (Fanuc)
      FLT_SyncPosition : Bool;   // Faulty snchronosation position
      FLT_1_1 : Bool;
      FLT_1_2 : Bool;
      FLT_1_3 : Bool;
      FLT_1_4 : Bool;
      FLT_1_5 : Bool;
      FLT_1_6 : Bool;
      FLT_1_7 : Bool;
      MSG_Rob_not_in_automatic : Bool;   // Interface in automatic but robot not in automatic
      MSG_Emergency_stop_Robot : Bool;   // Emergency stop robot
      MSG_2_2 : Bool;
      MSG_2_3 : Bool;
      MSG_2_4 : Bool;
      MSG_2_5 : Bool;
      MSG_2_6 : Bool;
      MSG_2_7 : Bool;
      MSG_3_0 : Bool;
      MSG_3_1 : Bool;
      MSG_3_2 : Bool;
      MSG_3_3 : Bool;
      MSG_3_4 : Bool;
      MSG_3_5 : Bool;
      MSG_3_6 : Bool;
      MSG_3_7 : Bool;
   END_STRUCT;
END_TYPE

TYPE "ABB_IRC6_State"
TITLE = Signals interface robot
VERSION : 0.0
   STRUCT
      Auto_mode_requested : Bool;   // Automatic mode requested
      Manual_mode_requested : Bool;   // Manual mode requested
      Auto_accepted : Bool;   // Automatic accepted
      Freigabe_Schaeumzyklus : Bool;   // Release foaming
      Release_foaming : Bool;   // Start foaming cycle
      Shot_time_received : Bool;   // Shot time received
      Data_transmitted : Bool;   // Data transmitted
      Data_inv_transmitted : Bool;   // Data inverse transmitted
      Interface_OK : Bool;   // Interface OK
      STG_System : Bool;   // Fault from system
      Fault_from_system : Bool;   // Fault from interface
      Fault_observed : Bool;   // Fault observed
      Escape_program : Bool;   // Escape program
      Motion_prog01_existing : Bool;   // Motion program 1 existing
      Motion_prog02_existing : Bool;   // Motion program 2 existing
      Motion_prog03_existing : Bool;   // Motion program 3 existing
      Robot_ProgNo_Mould_1 : Byte;   // Roboter program number mould 1
      Robot_ProgNo_Mould_2 : Byte;   // Roboter program number mould 2
      Robot_ProgNo_Mould_3 : Byte;   // Roboter program number mould 3
      Robot_processing_prog : Bool;   // Roboter processing program
      HFShotDigOut_open_MH : Bool;
      doShotDigOut_open_MH : Bool;
      HF_next_partshot : Bool;   // Flankenhilfsmerker für die Ermittlung eines neuen Verfahrprogramms // Teilschuß
      HF_Robot_not_in_Auto : Bool;   // Flankenhilfsmerker für das zurücksetzten des Signals "Roboter nicht in Auto"
      Robot_not_in_Auto : Bool;   // Roboter not in automatic mode
      Start_Synchronization : Bool;
      FLT_SyncPosition : Bool;   // Robot will perform the synchronization
      FHM_SyncEPS : Bool;   // The Synchronization position is not correct
      CleaningSelected : Bool;   // Flag for the information that a cleaning was selected
      CleaningActiv : Bool;   // Flag for the information that a cleaning is activ
      FHM_CleaningActiv : Bool;   // Helpflag for the information that a cleaning is activ
      FHM_start_test_shot : Bool;   // Flag for start test shot
      Start_test_shot : Bool;   // Start test shot with robot
      Reserve_6_6 : Bool;
      Reserve_6_7 : Bool;
      Reserve_7_0 : Bool;
      Reserve_7_1 : Bool;
      Reserve_7_2 : Bool;
      Reserve_7_3 : Bool;
      Reserve_7_4 : Bool;
      Reserve_7_5 : Bool;
      Reserve_7_6 : Bool;
      Reserve_7_7 : Bool;
      Reserve_Word_8 : Word;
      Reserve_Word_10 : Word;
      MC_Place_Number : Byte;
      Mould_Number : Byte;
      Time_Nummer : Byte;
      Offset_of_Shottime : Byte;
      Stepnumber : Byte;   // Schrittmerker für die Ablaufsteuerung der Roboteransteuerung
      Input : "ABB_IRC6_Input";   // Merkerbereich für die Eingänge vom Roboter
      Output : "ABB_IRC6_Output";   // Merkerbereich für die Ausgänge vom Roboter
      Meldungen : "ABB_IRC6_Messages";   // Merkerbereich für die Meldungen vom Roboter
   END_STRUCT;
END_TYPE

TYPE "IDM_115_FlowSpeedFloat"
VERSION : 0.1
   STRUCT
      Address : Hw_Io;
      Active : Bool;
      ChckConnFault : Bool;
      ChckConnDone : Bool;
      Skalierung : Struct
         Request : Bool;
         Transmitting : Bool;
         Active : Bool;
         Data : Struct
            Kalibrierfaktor : Real;
            Filterzeit : Word;
         END_STRUCT;
      END_STRUCT;
   END_STRUCT;
END_TYPE

TYPE "UDT702_HeatingControl"
TITLE = Parameter of tempering control (2 point)
VERSION : 0.1
   STRUCT
      Dif_Heating_ON : Real;   // Difference to switch the heating mode on
      Dif_Heating_OFF : Real;   // Difference to switch the heating mode on
      Max_Temp : Real;   // Max temperature to stop heating (absolute value)
   END_STRUCT;
END_TYPE

TYPE "UDT105_ControllerHeating"
TITLE = State of 2-point controller tempering
VERSION : 0.1
   STRUCT
      HeatingExists : Bool;
      HeatingActive : Bool;
      HeatingRequest : Bool;
      HeatingRelease : Bool;
      HF_Set_Cooling : Bool;
      HF_Set_Heating : Bool;
      HeatingExist : Bool;
      Fault_Exist : Bool;
      INFuse : Bool;
      INHeatingLimit : Bool;
      OUTHeating : Bool;
      Spare_1_6 : Bool;
      Spare_1_7 : Bool;
      Spare_1_8 : Bool;
      Spare_1_9 : Bool;
      Switch_ON_OFF : Bool;
      State_Temp : Int;
   END_STRUCT;
END_TYPE

TYPE "UDT754_Heating_State"
VERSION : 0.1
   STRUCT
      Supply_Heating_Exist : Array[1..1] of Bool;
      Exause_Heating_Exist : Array[1..1] of Bool;
      PreLIne_heating_Exist : Array[1..1] of Bool;
      ReturnLine_Heating_Exist : Array[1..1] of Bool;
   END_STRUCT;
END_TYPE

TYPE "ABB_IRC6_Input"
VERSION : 0.0
   STRUCT
      diMotorOn : Bool;   // Systeminput: Switch ON the motors of the robot
      diMotorOff : Bool;   // Systeminput: Switch OFF the motors of the robot
      diStartProg : Bool;   // Systeminput: Start the robotprogram from the last position in the program
      diStartMain : Bool;   // Systeminput: Start the robotprogram from the beginning
      diStopProg : Bool;   // Systeminput: Stop the robotprogram
      diResetError : Bool;   // Systeminput: Reset an systemerror
      diResetEstop : Bool;   // Systeminput: Reset the emergencystop
      diQuickStop : Bool;   // Systeminput: Stop the robot directly and switch the break ON
      diBreak : Bool;   // Signal to call the interrupt 1
      diInterrupt : Bool;   // Signal to call the interrupt 2
      diStartCycle : Bool;   // Signal to start the robotcycle
      diReadProgNo : Bool;   // A programnumber can read from PLC
      diStartMoveMC : Bool;   // The robot can start with it´s movements
      diShotDigIn : Bool;   // The foaming enabling of the machine is existing
      diStartBrushMH : Bool;   // Die Freigabe zum reinigen des MK's steht an (Bürstenstation ist bereit)
      diHomePrePos : Bool;   // Signal to move the robot from to the pre position
      diHomeToMaintP : Bool;   // Signal to move the robot from homeposition to maintenanceposition
      diMaintToHomeP : Bool;   // Signal to move the robot from maintenanceposition to homeposition
      diHomeToMaint2 : Bool;   // Signal to move the robot from homeposition to maintenanceposition 2
      diMaintToHome2 : Bool;   // Signal to move the robot from maintenanceposition 2 to homeposition
      diProgBreak : Bool;   // Signal to break the program
      di01_022 : Bool;   // Spare
      di01_023 : Bool;   // Spare
      di01_024 : Bool;   // Spare
      di01_025 : Bool;   // Spare
      di01_026 : Bool;   // Spare
      diRobinSavepos : Bool;   // Signal das der Weg in die Grund/ Wartungsposition frei ist
      diJumpConveyer : Bool;   // Signal to jump the routine "Conveyer- Tracking"
      diPLCWaitWobj : Bool;   // Signal to activate the waitwobj instruction
      diPLCDropWobj : Bool;   // Signal to drop the activ wobj
      diBackToRest : Bool;   // Signal to move the robot back to homeposition after foaming
      diStartEscape : Bool;   // Signal to move the robot to it´s escapeposition (anticollision)
      di01_033 : Bool;   // Spare
      diStartSyncSafety : Bool;   // Signal to move the robot to the syncronisation switch
      di01_035 : Bool;   // Spare
      di10_036 : Bool;   // Spare
      di10_037 : Bool;   // Spare
      di10_038 : Bool;   // Spare
      di10_039 : Bool;   // Spare
      di10_040 : Bool;   // Spare
      di10_041 : Bool;   // Spare
      diHomeToSprayP : Bool;   // Signal to move the robot to the Spray position
      diSprayToHomeP : Bool;   // Signal to move the robot to home position from spray position
      diRelSprayMould_1 : Bool;   // Release Release agent mould 1
      diRelSprayMould_2 : Bool;   // Release Release agent mould 2
      diRelSprayMould_3 : Bool;   // Release Release agent mould 3
      diRelSprayMould_4 : Bool;   // Release Release agent mould 4
      diRelFoamMould_1 : Bool;   // Release foaming mould 1
      diRelFoamMould_2 : Bool;   // Release foaming mould 2
      diRelFoamMould_3 : Bool;   // Release foaming mould 3
      diRelFoamMould_4 : Bool;   // Release foaming mould 4
      diCloseM_to_PP : Bool;
      diCloseM_to_EP : Bool;
      diCloseM_to_HP : Bool;
      di01_055 : Bool;   // Spare
      di01_056 : Bool;   // Spare
      di01_057 : Bool;   // Spare
      di01_058 : Bool;   // Spare
      di01_059 : Bool;   // Spare
      diStartCleanMH : Bool;   // The robot can move to MH-Cleaningstation
      diCleanMHEnd : Bool;   // The MH-Cleaning is finished
      di10_62 : Bool;   // Spare
      di10_63 : Bool;   // Spare
      di10_64 : Bool;   // Spare
      diStartFlushSpray : Bool;   // Signal that flushing started
      diEndFlushSpray : Bool;   // Signal flushing end
      diStartNextPart : Bool;   // Signal to enable the second partshot
      di01_068 : Bool;   // Spare
      di01_069 : Bool;   // Spare
      di01_070 : Bool;   // Spare
      di01_071 : Bool;   // Spare
      di01_072 : Bool;   // Spare
      di01_073 : Bool;   // Spare
      di01_074 : Bool;   // Spare
      di01_075 : Bool;   // Spare
      di01_076 : Bool;   // Spare
      di01_077 : Bool;   // Spare
      di01_078 : Bool;   // Spare
      di01_079 : Bool;   // Spare
      di01_080 : Bool;   // Spare
      giMouldCodeBit0 : Bool;   // Anzahl der Formen im Formträger (Gruppeingang Bit 0)
      giMouldCodeBit1 : Bool;   // Anzahl der Formen im Formträger (Gruppeingang Bit 1)
      giMouldCodeBit2 : Bool;   // Anzahl der Formen im Formträger (Gruppeingang Bit 2)
      di10_84 : Bool;   // Spare
      di10_85 : Bool;   // Spare
      di10_86 : Bool;   // Spare
      di10_87 : Bool;   // Spare
      di10_88 : Bool;   // Spare
      GIMCNo : Byte;   // Nummer des Formträgers der Form// Abhängig vom MouldCode
      GIProgNo1 : Word;   // Programnumber 1 (left mould in mould carrier)
      GIShotTX1 : Word;   // Schußzeit des nächsten Teilschusses in 1/10 Sekunden
   END_STRUCT;
END_TYPE

TYPE "ABB_IRC6_Output"